REGION Network 2: Select with vacuum
   VAK:  NOP   0;
         SET;
         =     #OUT_H_Vacuum_active;
   //
         AN    #IN_P_Vacuum;
         L     S5T#500MS;
         SD    #IN_Timer_delay_Lock;
   //
         A     #IN_P_Vacuum;
         L     S5T#500MS;
         SD    #IN_Timer_delay_Pumpe;
   //
         AN    #IN_P_Vacuum;
         A     #IN_Timer_delay_Lock;
         =     #OUT_V_Lock_Vacuum;
   //
         ON    #IN_P_Vacuum;
         ON    #IN_Timer_delay_Pumpe;
         =     #OUT_V_Pump_Vacuum;
   //
         L     1;
         T     #IO_Status.Status_Vacuum;
END_REGION
END_FUNCTION

FUNCTION "FC107_Binär->Bit" : Void   // FC107, STL
TITLE = Chang a bin value in a bitcodetd value
{ S7_Optimized_Access := 'FALSE' }
AUTHOR : KT242
FAMILY : RS_KK
NAME : BintoBit
VERSION : 1.0
   VAR_INPUT
      IN_BinaerZahl : Byte;   // Eingabe einer Zahl (Maximal 16) als Ganzzahl
   END_VAR
   VAR_OUTPUT
      OUT_BitZahl : Word;   // Ausgabe der Zahl als Bitcodiertes Word
   END_VAR
   VAR_TEMP
      Temp_Sprungzaehler : Word;   // Zwischenmerker für einen Schleifenzähler
      Temp_Out_BitZahl : Word;
   END_VAR
BEGIN

REGION Network 1
         L     0;
         T     #Temp_Out_BitZahl;
   //
         O(;
         L     16;
         L     #IN_BinaerZahl;
         <I;
         );
         O(;
         L     1;
         <I;
         );
         JC    ENDE;
   //
         L     1;
         T     #Temp_Out_BitZahl;
   //
         L     #IN_BinaerZahl;
         ==I;
         JC    ENDE;
         L     1;
         -I;
   //
   NEXT: NOP   0;
         T     #Temp_Sprungzaehler;
   //
         L     #Temp_Out_BitZahl;
         SLW   1;
         T     #Temp_Out_BitZahl;
   //
         L     #Temp_Sprungzaehler;
         LOOP  NEXT;
   ENDE: NOP   0;

         L     #Temp_Out_BitZahl;
         T     #OUT_BitZahl;
END_REGION
END_FUNCTION

FUNCTION "FC111_FIFO" : Void   // FC111, STL
TITLE = FIFO of interface numbers
{ S7_Optimized_Access := 'FALSE' }
AUTHOR : KT242
FAMILY : RS_KK
NAME : FIFO
VERSION : 1.0
   VAR_INPUT
      IN_Amount_Interfaces : Int;   // Amount of interfaces to start shotcycle
      IN_Register : "UDT001_DWord_1_32";   // Data area of registered interfaces
      IN_Reset_List : Bool;   // Reset of list by new start of plc
      IN_StartAdr : Pointer;   // Start-addresse at DB to save countervalues to find out position at FIFO
      IN_DataBlock : DB_ANY;   // Datablock to save countervalues to find out position at FIFO
   END_VAR
   VAR_IN_OUT
      IO_FIRST : Int;   // Number of the member at first positon
      IO_SECOND : Int;   // Number of the member at second positon
      IO_FlagNewPos : Bool;   // Flag determine new positions at fifo
   END_VAR
   VAR_TEMP
      Schleifengroesse : Int;   // Schleifenzähler für den Durchlauf der Positionen bis "IN_Anzahl_Teilnehmer"
      Aktueller_Wert : Word;   // Wert des Zähler der eingetragenen Schnittstelle zur Erkennung der Position
      Wert_First : Word;   // Wert des Zähler der am längsten (first) eingetragenen Schnittstelle
      Wert_Second : Word;   // Wert des Zähler der am nächsten (second) eingetragenen Schnittstelle
      Baustein_Nr : Int;   // Merker zur Erkennung des Speicherbereiches der Bits "IN_Eintragen"
      Adresse_im_Baustein : DWord;   // and the start adress within the program block
      Eintragen_lokal : DWord;   // Zwischenspeicher der eingetragenen Formträgerschnittstellen (von UDT auf DWORD)
   END_VAR
BEGIN

REGION Network 1: FIFO - buffer
   // Am Ausgang "FIRST" liegt die Nummer des ersteingetragenen und an "SECOND" die 
   // des nachfolgenden Teilnehmers (max. 16) an. 
   // Am Eingangswort "Eintragen" muß das entsprechende Bit solange TRUE sein, bis
   // der Teilnehmer wieder ausgetragen werden kann.
   // Das Austragen des Teilnehmers erfolgt, wenn sich dieser in der Position "FIRST" 
   // oder "SECOND" befindet, innerhalb des Bausteins für die Schnittstelle.
   //_______________________________________________________________
   // Schieben der Eingetragenen FTs auf lokalen DWord- Bereich
   //
         L;
         LAR1;
         L     W[AR1, P#0.0];
         T     #Baustein_Nr;
   //
         L     D[AR1, P#2.0];
         T     #Adresse_im_Baustein;
         LAR2;
         L;
         LAR1;
   //
         OPN   DB[ #Baustein_Nr];
         L     DBD[AR2, P#0.0];
         T     LD[AR1, P#0.0];
   //__________________________________________________________
   //
         L     0;
         T     #Schleifengroesse;
         T     #Wert_First;
         T     #Wert_Second;
         L;
         LAR2;
   //
         L     #Eintragen_lokal;
         CAD;
         T     #Eintragen_lokal;
   //
         L;
         LAR1;
   //
         A(;
         L     #Eintragen_lokal;
         L     0;
         <>D;
         );
         JC    NEXT;
   //
   NEXT: A     "Flag_02_500_Hertz";
         FP    #IO_FlagNewPos;
         JCN   ENDE;
   //
         L     0;
         T     #IO_FIRST;
         T     #IO_SECOND;
   //
   M002: A     [AR1, P#0.0];  // Eintragebit ist gesetzt
         JCN   M001;
   //
         OPN   #IN_DataBlock;
         L     DBW[AR2, P#0.0];  // Speicherwert für eingetragene Station
         +     1;  // um 1 erhöhen
         T     DBW[AR2, P#0.0];
         T     #Aktueller_Wert;
   //
         L     #Aktueller_Wert;  // Wenn Speicherwert grösser als Maximum ist
         L     #Wert_First;
         >I;
         JCN   M011;
   //
         L     #Wert_First;
         T     #Wert_Second;
   //
         L     #Aktueller_Wert;  // Speicherwert in Maximum übertragen
         T     #Wert_First;
   //
         L     #IO_FIRST;
         T     #IO_SECOND;
   //
         L     #Schleifengroesse;  // Nummer der ersteingetragenen Station
         +     1;
         T     #IO_FIRST;
   //
         JU    M001;
   //
   M011: NOP   0;
         L     #Aktueller_Wert;  // Wenn Speicherwert grösser als Maximum ist
         L     #Wert_Second;
         >I;
         JCN   M001;
   //
         L     #Aktueller_Wert;  // Speicherwert in Maximum übertragen
         T     #Wert_Second;
   //
         L     #Schleifengroesse;  // Nummer der ersteingetragenen Station
         +     1;
         T     #IO_SECOND;
   //
   M001: A     [AR1, P#0.0];  // Eintragebit ist gesetzt
         JC    M003;
         L     0;  // wenn nicht gesetzt, dann ablöschen
         OPN   #IN_DataBlock;
         T     DBW[AR2, P#0.0];
   //
   M003: L     #Schleifengroesse;
         +     1;
         T     #Schleifengroesse;  // nächste Station
         +AR1  P#0.1;
         +AR2  P#2.0;
         L     #Schleifengroesse;  // Schleife ausführen,
         L     #IN_Amount_Interfaces;  // bis zur Anzahl der Teilnehmer
         <I;
         JC    M002;
   //
   ENDE: NOP   0;
END_REGION
END_FUNCTION

FUNCTION "FC112_IF_SP_MC" : Void   // FC112, STL
TITLE = Interface to switch panel and mould carrier
{ S7_Optimized_Access := 'FALSE' }
AUTHOR : KT242
FAMILY : RS_KK
NAME : SS_FT
VERSION : 1.4
// Function block to book in interface-no. of a foaming cycle by operation panel 
// or mould carrier interface.
   VAR_INPUT
      IN_InterfaceNo : Int;   // Number of related Interface
      IN_PositionFIRST : Int;   // No of interface, which is at first position // from FC 111 FIFO
      IN_PositionSECOND : Int;   // No of interface, which is at second position // from FC 111 FIFO
      IN_BCDSwitchPrgrNo_MH : Byte;   // Inputbyte of program no. from program selection switch at mixinghead panel
      IN_MH_Automatic : Bool;   // Mode switch mixing head panel at position cycle start "Auto"
      IN_MH_Manual : Bool;   // Mode switch mixing head panel at position cycle start "Manual"
      IN_Start_MH_Panel : Bool;   // Button start cycle at mixing head panel to enter interface no. -> FIFO
      IN_Stop_MH_Panel : Bool;   // Button stop cycle at mixing head panel to erase interface no. -> FIFO
      IN_ResetFault : Bool;   // Quit fault within this function block
      IN_ReleaseSWU : Bool;   // Switch over unit (SWU) of this interface is released
      IN_ReleaseMouldcarrier : Bool;   // Foaming release of mouldcarrier to enter interface number -> FIFO
      IN_PrgNoSwitchDeselected : Bool;   // Signal to bridge program selection by program selection switch
      IN_ReleaseFoaming : Bool;   // External signal release entering interface number
      IN_ReleaseCycle : Bool;   // Release start foaming cycle from function block cycle is active
      IN_OperationModeAuto : Bool;   // Foaming machine in automatic mode
      IN_OperationModeTest : Bool;   // Foaming machine in test mode; no foaming over mixinghead
      IN_LampTest : Bool;   // Check indicator lamp selected
      IN_CycleRunning : Bool;   // Foaming cycle is active
      IN_ShotRunning : Bool;   // Foaming active
      IN_LastStandbyTimeCycle : Bool;   // Last shot of foaming cycle was carried out
      IN_PulseCycleFinished : Bool;   // Pulse foaming cycle finished
   END_VAR
   VAR_OUTPUT
      OUT_Fault_To_MC : Bool;   // Output fault happend at active interface
      OUT_ShotEnd_To_MC : Bool;   // Output all part shots finished at this interface
      OUT_H_MH_Panel : Bool;   // Indicator foaming release and state of foaming cycle at mixinghead panel
   END_VAR
   VAR_IN_OUT
      IO_InterfaceActiveFIFO : Bool;   // Information interface no. active at FIFO
      IO_Status : "UDT112_IF_UP_MC";
      IO_Fault : "UDT1816_FLT_IF_SP_MC";
      IO_NewFault : Bool;
      IO_FaultLevel_1 : Bool;
      IO_FaultLevel_3 : Bool;
   END_VAR
   VAR_TEMP
      Temp_IO_Status : "UDT112_IF_UP_MC";
      TEMP_IO_Fault : "UDT1816_FLT_IF_SP_MC";
      Temp_ERROR_CODE : Int;   // Error state of systemfunction "BLKMOV" Blockmove
      AnyPointer1 : ANY;   // Pointer to copy thr array "IO_Status" and "Temp_IO_Status"
      AnyPointer2 : ANY;   // Pointer to copy thr array "IO_Status" and "Temp_IO_Status"
      Temp_SelectionPrgNo_OK : Bool;   // Flag selction program no. is OK at mixing head panel
      Temp_Flag_RelInterface : Bool;   // Flag release interface to enter at FIFO
      Temp_Pulse_RelInterface : Bool;   // Pulse für enter interface no. at FIFO
      Temp_Interface_at_Pos_1 : Bool;   // Flag interface at first position at FIFO
      Temp_Interface_at_Pos_2 : Bool;   // Flag interface at second position at FIFO
      Temp_Interface_Deselect : Bool;   // Flag deselct interface at FIFO
      Temp_Value_1 : Word;   // Value to calculate view between FUP/ KOP
      Temp_Value_2 : Int;   // Value to calculate view between FUP/ KOP
   END_VAR
BEGIN

REGION Network 1: Saved data integration
   // Änderungen:
   // -------------------------------------------------------------------------------
   // Anpassung der Aufschlüsselung der Schnittstellenstörungen.
   // v.d.Geest     20.09.2005
   // -------------------------------------------------------------------------------
   // Bei einer Störung der Gruppe 1 oder bei den zurücknehmen der Schäumfreigabe 
   // wird nur noch die Schnittstelle an der Position 1 ausgetragen.
   // (Änderungen auch im UDT112)
   // v.d.Geest     29.11.2004
   // -------------------------------------------------------------------------------
   // Genauere Aufschlüsselung der Schnittstellenstörungen. (Änderungen auch im 
   // UDT112)
   // Lindner       12.07.2004
   // -------------------------------------------------------------------------------
   // Bei Anwahl der Betriebsart "Testen" wird die Anzeigen der Schäumfreigabe an dem 
   // Bedienpult nicht mehr angezeigt.
   // Bereits vor dem einschalten der Betriebsart "Testen" eingetragene 
   // Schnittstellen werden noch bearbeitet, es können aber keine neuen eingetragen 
   // werden.
   // v.d.Geest     08.04.2003
   // -------------------------------------------------------------------------------
   // Das Signal "OUT_Schussende_an_FT" wurde über das Signal nach Ablauf der 
   // Kreislaufzeit 2 gebildet. Hierdurch konnte es vorkommen das sich mehrere 
   // Formträger die sich zum Schäumen angemeldet haben innerhalb eines Ablaufs der 
   // KLZ 2 abmelden. (Änderungen auch im UDT112)
   // v.d.Geest     17.03.2003
   // -------------------------------------------------------------------------------
   //-----
         LAR1;
         L;
         LAR2;
   //-----
         L     16#1002;  // Bytes
         T     W[AR1, P#0.0];
         L     2;  // Amount of bytes
         T     W[AR1, P#2.0];
         L     W[AR2, P#0.0];  // Block no,
         T     W[AR1, P#4.0];
         L     D[AR2, P#2.0];  // Startadress of datas
         T     D[AR1, P#6.0];
   //-----
         CALL  BLKMOV
         ( SRCBLK  := #AnyPointer1,
           RET_VAL := #Temp_ERROR_CODE,
           DSTBLK  := #Temp_IO_Status
         );
   //-----
         LAR1;
         L;
         LAR2;
   //-----
         L     16#1002;  // Bytes
         T     W[AR1, P#0.0];
         L     2;  // Amount of bytes
         T     W[AR1, P#2.0];
         L     W[AR2, P#0.0];  // Block no,
         T     W[AR1, P#4.0];
         L     D[AR2, P#2.0];  // Startadress of datas
         T     D[AR1, P#6.0];
   //-----
         CALL  BLKMOV
         ( SRCBLK  := #AnyPointer2,
           RET_VAL := #Temp_ERROR_CODE,
           DSTBLK  := #TEMP_IO_Fault
         );
   //-----
END_REGION

REGION Network 2: Test the program / program no. OK
   // Eine Schäumfreigabe über diese Schnittstelle darf nur erfolgen, wenn die 
   // Programmvorwahl ok ist. Dieses ist im Handbetrieb der Fall, sobald eine gültige 
   // Programmnummer an dem Wahlschalter des Mischkopfbedienpultes eingestellt wurde.
   //-----
         A(;
         A(;
         A(;
         L     #IN_BCDSwitchPrgrNo_MH;
         T     #Temp_Value_1;
         SET;
         SAVE;
         CLR;
         A     BR;
         );
         JNB   _001;
         L     #Temp_Value_1;
         L     16#FF;
         AW;
         T     #Temp_Value_1;
         SET;
         SAVE;
         CLR;
   _001: A     BR;
         );
         JNB   _002;
         L     #Temp_Value_1;
         T     #Temp_Value_2;
         SET;
         SAVE;
         CLR;
   _002: A     BR;
         );
         A(;
         L     #Temp_Value_2;
         L     0;
         <>I;
         );
         O     #IN_PrgNoSwitchDeselected;
         O(;
         A     #IN_CycleRunning;
         AN    #IN_Start_MH_Panel;
         AN    #IN_LastStandbyTimeCycle;
         );
         =     #Temp_SelectionPrgNo_OK;
END_REGION

REGION Network 3: Interface at position 1 of FIFO
         L     #IN_PositionFIRST;
         L     #IN_InterfaceNo;
         ==I;
         =     #Temp_IO_Status.IF_is_on_1_Position;
         =     #Temp_Interface_at_Pos_1;
END_REGION

REGION Network 4: Interface number to start next
         L     #IN_PositionSECOND;
         L     #IN_InterfaceNo;
         ==I;
         =     #Temp_IO_Status.IF_is_on_2_Position;
         =     #Temp_Interface_at_Pos_2;
END_REGION

REGION Network 5: Release mould carrier
         A(;
         A     #IN_MH_Automatic;
         A     #IN_ReleaseMouldcarrier;
         O     #IN_MH_Manual;
         );
         A     #Temp_SelectionPrgNo_OK;
         =     #Temp_Flag_RelInterface;
END_REGION

REGION Network 6: Sign out mouldcarrier by button Stop- foaming
         AN    #Temp_Interface_at_Pos_1;
         AN    #Temp_Interface_at_Pos_2;
         AN    #IN_Stop_MH_Panel;
         A     #IN_MH_Manual;
         S     #Temp_IO_Status.Stop_Buton_switched;
         A(;
         A     #IN_MH_Manual;
         A     #IN_Start_MH_Panel;
         A     #Temp_IO_Status.Stop_Buton_switched;
         ON    #Temp_IO_Status.IF_is_Selected;
         );
         R     #Temp_IO_Status.Stop_Buton_switched;
         NOP   0;
END_REGION

REGION Network 7: Fault at the interface
         A(;
         A(;
         ON    #IN_MH_Automatic;
         O     #IN_ResetFault;
         );
         R     #TEMP_IO_Fault.Fault_IF;

         A(;
         AN    #IN_MH_Manual;
         AN    #IN_MH_Automatic;
         O(;
         AN    #Temp_Flag_RelInterface;
         A     #IN_CycleRunning;
         AN    #IN_LastStandbyTimeCycle;
         );
         O(;
         A(;
         O     #IO_FaultLevel_1;
         ON    #IN_ReleaseFoaming;
         ON    #IN_ReleaseCycle;
         );
         FP    #Temp_IO_Status.FHF_Fault;
         AN    #IN_LastStandbyTimeCycle;
         A     #Temp_Interface_at_Pos_1;
         );
         ON    #IN_OperationModeAuto;
         ON    #IN_ReleaseSWU;
         O;
         A(;
         O     #Temp_Interface_at_Pos_1;
         O     #Temp_Interface_at_Pos_2;
         );
         A(;
         O     #Temp_IO_Status.Stop_Buton_switched;
         ON    #IN_Stop_MH_Panel;
         );
         );
         A     #Temp_IO_Status.IF_is_Selected;
         AN    #TEMP_IO_Fault.Fault_IF;
         S     #IO_NewFault;
         S     #TEMP_IO_Fault.Fault_IF;
         A     #TEMP_IO_Fault.Fault_IF;
         );
         A     #IN_MH_Automatic;
         =     #OUT_Fault_To_MC;
END_REGION

REGION Network 8: Shotend
         A(;
         A(;
         ON    #IN_MH_Automatic;
         O;
         AN    #Temp_Flag_RelInterface;
         AN    #TEMP_IO_Fault.Fault_IF;
         );
         R     #Temp_IO_Status.Shotsend_IF;
         A(;
         O     #TEMP_IO_Fault.Fault_IF;
         O     #IN_PulseCycleFinished;
         );
         FP    #Temp_IO_Status.FHF_KLZ2;
         A     #Temp_Interface_at_Pos_1;
         S     #Temp_IO_Status.Shotsend_IF;
         A     #Temp_IO_Status.Shotsend_IF;
         );
         A     #IN_MH_Automatic;
         =     #OUT_ShotEnd_To_MC;
END_REGION

REGION Network 9: Log in interface no at FIFO
         A(;
         A     #IN_Start_MH_Panel;
         FP    #Temp_IO_Status.HF_T_Start_MH;
         A     #IN_MH_Manual;
         O;
         A(;
         A     #IN_ReleaseMouldcarrier;
         BLD   100;
         FP    #Temp_IO_Status.HF_Release_IF;
         );
         A     #IN_MH_Automatic;
         );
         AN    #IN_OperationModeTest;
         A     #Temp_Flag_RelInterface;
         A     #IN_ReleaseSWU;
         A     #IN_ReleaseFoaming;
         A     #IN_ReleaseCycle;
         AN    #Temp_IO_Status.IF_is_Selected;
         AN    #Temp_IO_Status.Shotsend_IF;
         AN    #TEMP_IO_Fault.Fault_IF;
         S     #Temp_IO_Status.IF_is_Selected;
         S     #IO_InterfaceActiveFIFO;
END_REGION

REGION Network 10: Log off interface no. at FIFO
         A     #IN_PulseCycleFinished;
         A     #Temp_Interface_at_Pos_1;
         O;
         AN    #Temp_Flag_RelInterface;
         AN    #Temp_Interface_at_Pos_1;
         ON    #IN_OperationModeAuto;
         O     #TEMP_IO_Fault.Fault_IF;
         A     #Temp_IO_Status.IF_is_Selected;
         =     #Temp_Interface_Deselect;
         R     #Temp_IO_Status.IF_is_Selected;
         R     #IO_InterfaceActiveFIFO;
END_REGION

REGION Network 11: Start cycle with this interface
         A     #Temp_IO_Status.IF_is_Selected;
         A     #Temp_Interface_at_Pos_1;
         A     #IN_ReleaseFoaming;
         A     #IN_ReleaseCycle;
         AN    #IN_CycleRunning;
         =     #Temp_IO_Status.Start_to_Cycle;
END_REGION

REGION Network 12: Break cycle at this interface
         AN    #Temp_IO_Status.IF_is_Selected;
         A     #Temp_Interface_at_Pos_1;
         AN    #IN_LastStandbyTimeCycle;
         A     #IN_CycleRunning;
         =     #Temp_IO_Status.Stop_to_Cycle;
END_REGION

REGION Network 13: Set indicater ready for foaming
         A(;
         A     #Temp_Flag_RelInterface;
         A     #IN_MH_Manual;
         O     #IN_MH_Automatic;
         );
         A     #IN_ReleaseFoaming;
         A     #IN_ReleaseCycle;
         A(;
         ON    #Temp_IO_Status.Shotsend_IF;
         O;
         A     #IN_LastStandbyTimeCycle;
         A     #Temp_Interface_at_Pos_1;
         );
         A(;
         AN    #Temp_IO_Status.IF_is_Selected;
         A     #IN_MH_Manual;
         AN    #IN_OperationModeTest;
         O;
         A     #Temp_IO_Status.IF_is_Selected;
         A(;
         AN    #Temp_Interface_at_Pos_1;
         A     "Flag_00_500_Hertz";
         O;
         A     #Temp_Interface_at_Pos_1;
         A(;
         AN    #IN_ShotRunning;
         A     "Flag_01_000_Hertz";
         O;
         A     #IN_ShotRunning;
         A     "Flag_05_000_Hertz";
         );
         );
         );
         A     #Temp_SelectionPrgNo_OK;
         A     #IN_ReleaseSWU;
         AN    #TEMP_IO_Fault.Fault_IF;
         O     #IN_LampTest;
         =     #OUT_H_MH_Panel;
END_REGION

REGION Network 14: Reset of faults
         O     #IN_ResetFault;
         R     #TEMP_IO_Fault.FLT_pouring_release;
         R     #TEMP_IO_Fault.FLT_SWU_release;
         R     #TEMP_IO_Fault.FLT_Stop_while_selected;
         R     #TEMP_IO_Fault.FLT_op_mode_O;
         R     #TEMP_IO_Fault.FLT_Cycle_release;
END_REGION

REGION Network 15: Fault foaming release (external signal)
   // Störung: Die Schäumfreigebe wurde auf 0 gesetzt. Während der Formträger 
   // angemeldet und an erster Position ist.
   // - #Temp_IO_Status.Stoerung_Schaeumfreigabe -
         AN    #IN_ReleaseFoaming;
         AN    #IN_LastStandbyTimeCycle;
         A     #Temp_Interface_Deselect;
         A     #Temp_Interface_at_Pos_1;
         A     #IN_MH_Automatic;
         AN    #TEMP_IO_Fault.FLT_pouring_release;
         S     #IO_NewFault;
         S     #TEMP_IO_Fault.FLT_pouring_release;
END_REGION

REGION Network 16: Fault SWU release set to 0 (external signal)
   // Störung: Die USE-Freigabe wurde auf 0 gesetzt. Während der Formträger 
   // angemeldet ist.
   // - #Temp_IO_Status.USE_Freigabe-
         AN    #IN_ReleaseSWU;
         A     #Temp_Interface_Deselect;
         AN    #TEMP_IO_Fault.FLT_pouring_release;
         AN    #TEMP_IO_Fault.FLT_SWU_release;
         S     #IO_NewFault;
         S     #TEMP_IO_Fault.FLT_SWU_release;
END_REGION

REGION Network 17: Fault STOP-button pressed during foaming cycle
   // Störung: Der STOP-Taster wurde auf 0 gesetzt. Während der Formträger 
   // angemeldet und an erster Position ist.
   // -#Temp_IO_Status.Stoerung_STOP_Taster-
         A(;
         O     #Temp_Interface_at_Pos_1;
         O     #Temp_Interface_at_Pos_2;
         );
         A(;
         O     #Temp_IO_Status.Stop_Buton_switched;
         ON    #IN_Stop_MH_Panel;
         );
         A     #Temp_Interface_Deselect;
         AN    #TEMP_IO_Fault.FLT_pouring_release;
         AN    #TEMP_IO_Fault.FLT_SWU_release;
         AN    #TEMP_IO_Fault.FLT_Stop_while_selected;
         S     #IO_NewFault;
         S     #TEMP_IO_Fault.FLT_Stop_while_selected;
END_REGION

REGION Network 18: Fault key-switch manual/auto at MH-panel set to 0
   // Störung: Der Hand/Auto Schlüsselschalter wurde auf 0 gesetzt. Während der 
   // Formträger angemeldet und an erster Position ist.
   // -#Temp_IO_Status.Stoerung_Hand_Auto-
         AN    #IN_MH_Manual;
         AN    #IN_MH_Automatic;
         A     #Temp_Interface_at_Pos_1;
         AN    #TEMP_IO_Fault.FLT_pouring_release;
         AN    #TEMP_IO_Fault.FLT_SWU_release;
         AN    #TEMP_IO_Fault.FLT_Stop_while_selected;
         AN    #TEMP_IO_Fault.FLT_op_mode_O;
         S     #IO_NewFault;
         S     #TEMP_IO_Fault.FLT_op_mode_O;
END_REGION

REGION Network 19: Fault foaming release
   // Störung: Freigabe Zyklus wurde auf 0 gesetzt. Während der 
   // Formträger angemeldet und an erster Position ist.
         AN    #IN_ReleaseCycle;
         AN    #IN_LastStandbyTimeCycle;
         A     #Temp_Interface_at_Pos_1;
         AN    #TEMP_IO_Fault.FLT_pouring_release;
         AN    #TEMP_IO_Fault.FLT_SWU_release;
         AN    #TEMP_IO_Fault.FLT_Stop_while_selected;
         AN    #TEMP_IO_Fault.FLT_op_mode_O;
         AN    #TEMP_IO_Fault.FLT_Cycle_release;
         S     #IO_NewFault;
         S     #TEMP_IO_Fault.FLT_Cycle_release;
END_REGION

REGION Network 20: Error handling
         O     #TEMP_IO_Fault.FLT_pouring_release;
         O     #TEMP_IO_Fault.FLT_SWU_release;
         O     #TEMP_IO_Fault.FLT_Stop_while_selected;
         O     #TEMP_IO_Fault.FLT_op_mode_O;
         O     #TEMP_IO_Fault.FLT_Cycle_release;
         O     #TEMP_IO_Fault.Fault_IF;
         S     #IO_FaultLevel_3;
END_REGION

REGION Network 21: Save data
   //-----
         CALL  BLKMOV
         ( SRCBLK  := #Temp_IO_Status,
           RET_VAL := #Temp_ERROR_CODE,
           DSTBLK  := #AnyPointer1
         );
   //-----
         CALL  BLKMOV
         ( SRCBLK  := #TEMP_IO_Fault,
           RET_VAL := #Temp_ERROR_CODE,
           DSTBLK  := #AnyPointer2
         );
   //-----
END_REGION
END_FUNCTION

FUNCTION "FC114_IF_externalPlant" : Void   // FC114, STL
TITLE = Interface between machine and external plant
{ S7_Optimized_Access := 'FALSE' }
AUTHOR : KT242
NAME : SS_AP
VERSION : 1.1
   VAR_INPUT
      IN_Release : Bool;   // General release of interface external plant
      IN_use_Inv_Program : Bool;   // Number transfer by using an inverse program number
      IN_use_Parity_Bit : Bool;   // Number transfer by using parity check
      IN_Reset_fault_Fkt : Bool;   // Signal to reset faults at innerhalb this function block
      IN_Stop_MH_OpPanel : Bool;   // Stop- signal at MH - operator panel to put out interfacenumber from FIFO
      IN_Operationmode_Operate : Bool;   // Foaming machine in operation mode with foam dispersion
      IN_MH_panel_automatic : Bool;   // Mixinghead - operator panel switched to automatic
      IN_FCycleRelease_extern : Bool;   // Foaming release from externen plant
      IN_FCycle_release : Bool;   // Release start foaming cycle from function block cycle
      IN_FCycle_running : Bool;   // Foaming cycle is running
      IN_FCycle_Shotrelease : Bool;   // Foaming release from Schäumzyklus steht an
      IN_FCycle_Shot_running : Bool;   // Foaming happens
      IN_FCycle_Pulse_Shotend : Bool;   // Foaming finished
      IN_FCycle_Pulse_End : Bool;   // Pulse foaming cycle finished // Signal takes 1 SPS- Cycle
      IN_ExtPlant_OK : Bool;   // Signal from external plant: External plant is ready for production
      IN_Strobe_or_Start : Bool;   // Signal from external plant: Strobe valid or cycle start signal
      IN_StrobeINV_or_Parity : Bool;   // Signal from external plant: Data strobe inverse or parity bit
      IN_Start_Shot : Bool;   // Signal from external plant: Start foaming by shot release from PU
      IN_CP_forward : Bool;   // Signal from external plant: Trigger cleaning piston
      IN_ProgNo_ExtPlant : Byte;   // Signal from external plant: Program no or inverse program number
      IN_maxAmount_ProgNo : Int;   // Limitation of program number from external plant
   END_VAR
   VAR_OUTPUT
      OUT_PU_OK : Bool;   // Signal to external Plant: Foaming machine is ready to start foaming cycle
      OUT_Strobe_quit : Bool;   // Signal to external Plant: Program number (..Invers) was accepted
      OUT_FCycle_running : Bool;   // Signal to external Plant: Foaming cycle was started and runs
      OUT_ReadyForFoaming : Bool;   // Signal to external Plant: Foaming machine ready to open mixinghead
      OUT_FoamingActive : Bool;   // Signal to external Plant: Foaming is going on
      OUT_FoamingEnd : Bool;   // Signal to external Plant: Foaming is finished
      OUT_ServiceShot : Bool;   // Signal to external Plant: Foaming machine is at service mode
   END_VAR
   VAR_IN_OUT
      IO_Status : "UDT114_IF_externalPlant";
      IO_Fault : "UDT1817_FLT_IF_extPlant";
      IO_NewFault : Bool;
      IO_FaultLevel_1 : Bool;
      IO_FaultLevel_2 : Bool;
      IO_FaultLevel_3 : Bool;
   END_VAR
   VAR_TEMP
      Temp_IO_Status : "UDT114_IF_externalPlant";
      TEMP_IO_Fault : "UDT1817_FLT_IF_extPlant";
      ERROR_CODE : Int;   // Error state of systemfunction "BLKMOV" Blockmove
      AnyPointer1 : ANY;   // Pointer to copy thr array "IO_Status" and "Temp_IO_Status"
      AnyPointer2 : ANY;   // Pointer to copy thr array "IO_Status" and "Temp_IO_Status"
      Temp_ProgNo_Puls : Byte;   // Temporärer Zwischenspeicher der Programmnummer für die Paritätsprüfung
      Strobe_quitt_reset : Bool;   // Hilfsmerker zum zurücksetzen des Quittierungsbits
      Temp_PulseCycleRelease : Bool;   // Impulshilfsmerker das das starten einen Schäumzyklusses Freigegeben ist
      Temp_Pulse_ExtP_Start : Bool;   // Impulshilfsmerker für das Starten die Programmermittlung des Schnittstelle
   END_VAR
BEGIN

REGION Network 1: Saved data integration
   // Änderungen:
   // -------------------------------------------------------------------------------
   // Wenn beim starten der Anlage das Stobe Bit von der Fremdanlage schon oder noch 
   // gesetzt war wurde direkt ein Schäumprogramm gestartet.
   // Durch eine Flankenabfrage des Signals "#IN_Strobe_oder_Start" im Netzwerk 3 
   // wurde dieses unterbunden
   // 
   // Jäger       19.08.2004
   // -------------------------------------------------------------------------------
   //-----
         LAR1;
         L;
         LAR2;
   //-----
         L     16#1002;  // Bytes
         T     W[AR1, P#0.0];
         L     6;  // Amount of bytes
         T     W[AR1, P#2.0];
         L     W[AR2, P#0.0];  // Block no,
         T     W[AR1, P#4.0];
         L     D[AR2, P#2.0];  // Startadress of datas
         T     D[AR1, P#6.0];
   //-----
         CALL  BLKMOV
         ( SRCBLK  := #AnyPointer1,
           RET_VAL := #ERROR_CODE,
           DSTBLK  := #Temp_IO_Status
         );
   //-----
         LAR1;
         L;
         LAR2;
   //-----
         L     16#1002;  // Bytes
         T     W[AR1, P#0.0];
         L     2;  // Amount of bytes
         T     W[AR1, P#2.0];
         L     W[AR2, P#0.0];  // Block no,
         T     W[AR1, P#4.0];
         L     D[AR2, P#2.0];  // Startadress of datas
         T     D[AR1, P#6.0];
   //-----
         CALL  BLKMOV
         ( SRCBLK  := #AnyPointer2,
           RET_VAL := #ERROR_CODE,
           DSTBLK  := #TEMP_IO_Fault
         );
   //-----
END_REGION

REGION Network 2: Reset and set of faults
         CLR;
         =     #Temp_IO_Status.FaultLevel_1;
         =     #Temp_IO_Status.FaultLevel_2;
         =     #Temp_IO_Status.FaultLevel_3;
         =     #Temp_IO_Status.Message_activ;
   //-----
         A     #IN_Reset_fault_Fkt;
         R     #TEMP_IO_Fault.FLT_Strobe;
         R     #TEMP_IO_Fault.FLT_Strobe_inv;
         R     #TEMP_IO_Fault.FLT_AP_not_OK;
         R     #TEMP_IO_Fault.FLT_no_number;
         R     #TEMP_IO_Fault.FLT_inverse_number;
         R     #TEMP_IO_Fault.FLT_Parity_Bit;
         R     #TEMP_IO_Fault.FLT_Cycle_Stoped;
         R     #TEMP_IO_Fault.FLT_Start_Shot;
   //
         O     #IN_FCycle_release;
         FP    #Temp_IO_Status.FHF_Cycle_Release;
         =     #Temp_PulseCycleRelease;
   //
         O     #Temp_PulseCycleRelease;
         ON    #IN_ExtPlant_OK;
         A     #IN_Strobe_or_Start;
         A     #IN_MH_panel_automatic;
         AN    #TEMP_IO_Fault.FLT_Start_Shot;
         AN    #TEMP_IO_Fault.FLT_no_number;
         AN    #TEMP_IO_Fault.FLT_Strobe;
         S     #TEMP_IO_Fault.FLT_Strobe;
         S     #IO_NewFault;
   //
         O     #Temp_PulseCycleRelease;
         ON    #IN_ExtPlant_OK;
         A     #IN_StrobeINV_or_Parity;
         AN    #IN_use_Parity_Bit;
         A     #IN_MH_panel_automatic;
         AN    #TEMP_IO_Fault.FLT_no_number;
         AN    #TEMP_IO_Fault.FLT_Strobe_inv;
         S     #TEMP_IO_Fault.FLT_Strobe_inv;
         S     #IO_NewFault;
   //
         A     #IN_ExtPlant_OK;
         A     #IN_FCycle_release;
         A     #IN_Start_Shot;
         A     #IN_Strobe_or_Start;
         A     #IN_MH_panel_automatic;
         AN    #Temp_IO_Status.PU_Shotend;
         AN    #Temp_IO_Status.IF_is_selected;
         AN    #TEMP_IO_Fault.FLT_Start_Shot;
         S     #TEMP_IO_Fault.FLT_Start_Shot;
         S     #IO_NewFault;
   //
         AN    #IN_ExtPlant_OK;
         A     #IN_Release;
         A     #IN_MH_panel_automatic;
         AN    #TEMP_IO_Fault.FLT_AP_not_OK;
         =     #TEMP_IO_Fault.MSG_AP_not_OK;
         S     #Temp_IO_Status.Message_activ;
   //
         AN    #IN_ExtPlant_OK;
         A     #IN_Release;
         A     #IN_FCycle_release;
         A     #IN_MH_panel_automatic;
         AN    #TEMP_IO_Fault.FLT_AP_not_OK;
         S     #TEMP_IO_Fault.FLT_AP_not_OK;
         S     #IO_NewFault;
   //
END_REGION

REGION Network 3: Raising edge of Start/ Strobe- signal
         A     #IN_Strobe_or_Start;
         FP    #Temp_IO_Status.HF_StrobeStart;
         =     #Temp_Pulse_ExtP_Start;
END_REGION

REGION Network 4: Release start signal detection
         A     #IN_FCycle_release;
         A     #IN_Release;
         A     #IN_ExtPlant_OK;
         A     #IN_Stop_MH_OpPanel;
         A     #IN_MH_panel_automatic;
         AN    #TEMP_IO_Fault.FLT_Strobe;
         AN    #TEMP_IO_Fault.FLT_Strobe_inv;
         AN    #TEMP_IO_Fault.FLT_Start_Shot;
         AN    #TEMP_IO_Fault.FLT_AP_not_OK;
         AN    #TEMP_IO_Fault.FLT_Parity_Bit;
         AN    #TEMP_IO_Fault.FLT_Cycle_Stoped;
         JCN   res;
END_REGION

REGION Network 5: Select signal transver mode (Invers or Parity)
   // Dieser Baustein kann wahlweise für verschiedene Fremdanlagenschnittstellen 
   // verwendet werden.
   // - Hardwareschnittstelle mit Programm und invertiertem Programm
   // - Profibusschnittstelle nur mit einer Programmnummer
   // - Schnittstelle mit Paritätsbitüberbrüfung
         A     #IN_use_Parity_Bit;
         JC    PaCh;  // Jump to parity check
END_REGION

REGION Network 6: Sprungleiste fuer Invers check
         L     #Temp_IO_Status."Step";
         JL    res1;
         JU    stro;  // case 0     Strobe
         JU    qstr;  // case 1     quitt Strobe
         JU    istr;  // case 2     Strobe invers
         JU    qist;  // case 3     quitt Strobe invers
         JU    wait;  // case 4     Wait till Null
   //
   res1: JU    res;
END_REGION

REGION Network 7: Strobe
   stro: NOP   0;
         A     #Temp_Pulse_ExtP_Start;  //Edge Strobe or Start signal
         JCN   ausg;
   //
         A(;
         L     #IN_ProgNo_ExtPlant;
         L     0;
         <=I;
         );
         A(;
         L     #IN_ProgNo_ExtPlant;
         L     #IN_maxAmount_ProgNo;
         >I;
         );
         AN    #TEMP_IO_Fault.FLT_no_number;
         S     #TEMP_IO_Fault.FLT_no_number;
         S     #IO_NewFault;
   //
         L     #IN_ProgNo_ExtPlant;
         T     #Temp_IO_Status.PrgNo_Storage;
   //
         A     #IN_use_Inv_Program;
         JC    J_qu;
   //
         L     3;
         T     #Temp_IO_Status."Step";
         JU    ausg;
   //
   J_qu: L     1;
         T     #Temp_IO_Status."Step";
   //
         JU    ausg;
END_REGION

REGION Network 8: Confirme strobe
   qstr: NOP   0;  // case 1
         A     #IN_Strobe_or_Start;
         S     #OUT_Strobe_quit;
   //
         AN    #IN_Strobe_or_Start;
         A     #OUT_Strobe_quit;
         R     #OUT_Strobe_quit;
         JCN   ausg;
         L     2;
         T     #Temp_IO_Status."Step";
         JU    ausg;
END_REGION

REGION Network 9: Strobe invers und check ob ok
   istr: NOP   0;  // case 2
         A     #IN_StrobeINV_or_Parity;
         JCN   ausg;
         L     #IN_ProgNo_ExtPlant;
         L     #Temp_IO_Status.PrgNo_Storage;
         +I;
         L     255;
         ==I;
         NOT;
         AN    #TEMP_IO_Fault.FLT_inverse_number;
         S     #TEMP_IO_Fault.FLT_inverse_number;
         S     #IO_NewFault;
   //
         L     3;
         T     #Temp_IO_Status."Step";
   //
         JU    ausg;
END_REGION

REGION Network 10: Confirm (Quitt) strobe invers
   qist: NOP   0;  // case 3
   //
         A     #IN_StrobeINV_or_Parity;
         A     #IN_use_Inv_Program;
         O     #IN_Strobe_or_Start;
         S     #OUT_Strobe_quit;
   //
         L     4;
         T     #Temp_IO_Status."Step";
   //
         AN    #TEMP_IO_Fault.FLT_no_number;
         AN    #TEMP_IO_Fault.FLT_inverse_number;
         S     #Temp_IO_Status.IF_is_selected;
   //
         JU    ausg;
END_REGION

REGION Network 11: Warte auf strobe/ strobe invers auf Null
   wait: NOP   0;  // case 4
   //
         A     #IN_StrobeINV_or_Parity;
         A     #IN_use_Inv_Program;
         O     #IN_Strobe_or_Start;
         JC    Next;
         L     0;
         T     #Temp_IO_Status."Step";
         SET;
         R     #OUT_Strobe_quit;
   //
   Next: NOP   0;
   //
         JU    ausg;  // Jump over Parity check
END_REGION

REGION Network 12: Parity Check
   PaCh: NOP   0;
   //
         A     #Temp_Pulse_ExtP_Start;
         AN    #Temp_IO_Status.IF_is_selected;
         JCN   ausg;
   //
         L     #IN_ProgNo_ExtPlant;
         T     #Temp_ProgNo_Puls;
         T     #Temp_IO_Status.PrgNo_Storage;
   //
         X     #Temp_ProgNo_Puls.%X0;
         X     #Temp_ProgNo_Puls.%X1;
         X     #Temp_ProgNo_Puls.%X2;
         X     #Temp_ProgNo_Puls.%X3;
         X     #Temp_ProgNo_Puls.%X4;
         X     #Temp_ProgNo_Puls.%X5;
         X     #Temp_ProgNo_Puls.%X6;
         X     #Temp_ProgNo_Puls.%X7;
         X     #IN_StrobeINV_or_Parity;
         S     #TEMP_IO_Fault.FLT_Parity_Bit;
         S     #IO_NewFault;

   //
         O(;
         L     0;
         L     #Temp_ProgNo_Puls;
         >=I;
         );
         O(;
         L     #IN_maxAmount_ProgNo;
         >I;
         );
         S     #TEMP_IO_Fault.FLT_no_number;
         S     #IO_NewFault;
   //
         AN    #TEMP_IO_Fault.FLT_Parity_Bit;
         AN    #TEMP_IO_Fault.FLT_no_number;
         S     #Temp_IO_Status.IF_is_selected;
   //
         JU    ausg;
END_REGION

REGION Network 13: Reset
   res:  NOP   0;
         A     #Temp_IO_Status.IF_is_selected;
         =     #Temp_IO_Status.Stop_to_Cycle;
   //     UN    #TEMP_IO_Fault.FLT_Cycle_Stoped
   //      S     #TEMP_IO_Fault.FLT_Cycle_Stoped
   //      S     #IO_NewFault
   //
         SET;
         R     #Temp_IO_Status.IF_is_selected;
         R     #OUT_Strobe_quit;
         R     #Temp_IO_Status.Start_to_Cycle;
         R     #Temp_IO_Status.ExtP_MH_open;
         R     #Temp_IO_Status.ExtP_CP_forward;
   //
         A     #IN_StrobeINV_or_Parity;
         O     #IN_Strobe_or_Start;
         =     #OUT_Strobe_quit;
   //
         L     0;
         T     #Temp_IO_Status."Step";
         T     #Temp_IO_Status.PrgNo_Storage;
END_REGION

REGION Network 14: Starten des Schäumzyklusses
   ausg: NOP   0;
   //
         A     #Temp_IO_Status.IF_is_selected;
         AN    #IN_FCycle_running;
         =     #Temp_IO_Status.Start_to_Cycle;
         JCN   shot;
   //
         L     #Temp_IO_Status.PrgNo_Storage;
         T     #Temp_IO_Status.PrgNo_to_PU;
   //
   shot: NOP   0;
   //
         O     #IN_FCycle_Pulse_End;
         JCN   Goon;
   //
         SET;
         R     #Temp_IO_Status.IF_is_selected;
         L     0;
         T     #Temp_IO_Status.PrgNo_to_PU;
   //
   Goon: NOP   0;
END_REGION

REGION Network 15: Bilden der Signale an die/ von der Fremdanlage
   //______________________________________________
   // Die Schäummaschine ist Betriebsbereit
   //
         A     #IN_Release;
         A     #IN_FCycle_release;
         A     #IN_MH_panel_automatic;
         =     #Temp_IO_Status.PU_ok;
   //
         A     #IN_FCycle_running;
         A     #IN_MH_panel_automatic;
         =     #Temp_IO_Status.PU_Cycle_runs;
   //______________________________________________
   // Freigabe zum Ansteuern des Mischkofes
   //
         A     #IN_FCycle_Shotrelease;
         AN    #Temp_IO_Status.PU_Shotend;
         =     #Temp_IO_Status.PU_Pouringrelease;
   //______________________________________________
   // Bilden des Signal Schuss beendet
   //
         A     #IN_FCycle_Pulse_Shotend;
         S     #Temp_IO_Status.PU_Shotend;
   //
         AN    #IN_Start_Shot;
         A     #Temp_IO_Status.PU_Shotend;
         S     #Temp_IO_Status.StatShotOffafterCycleFinish;
         AN    #IN_FCycle_running;
         A     #Temp_IO_Status.PU_Shotend;
         S     #Temp_IO_Status.CycleOffafterShotFinish;
   //
         A     #Temp_IO_Status.StatShotOffafterCycleFinish;
         A     #Temp_IO_Status.CycleOffafterShotFinish;
         R     #Temp_IO_Status.PU_Shotend;
         R     #Temp_IO_Status.StatShotOffafterCycleFinish;
         R     #Temp_IO_Status.CycleOffafterShotFinish;
   //______________________________________________
   // Ansteuern des Mischkopfventils von der Fremdanlage
   //
         A     #IN_Start_Shot;
         A     #IN_FCycle_running;
         A     #IN_MH_panel_automatic;
         AN    #Temp_IO_Status.PU_Shotend;
         =     #Temp_IO_Status.ExtP_MH_open;
   //______________________________________________
   // Ansteuern des Reinigungskolben von der Fremdanlage
   //
         A     #IN_CP_forward;
         =     #Temp_IO_Status.ExtP_CP_forward;
   //______________________________________________
   // Signal das sich die Fremdanlage im Automatikbetrieb befindet
   //
         A     #IN_ExtPlant_OK;
         =     #Temp_IO_Status.ExtP_in_Automatic;
END_REGION

REGION Network 16: Ansteuern der Signale an die Fremdanlage
         A     #Temp_IO_Status.PU_ok;
         =     #OUT_PU_OK;
   //
         A     #Temp_IO_Status.PU_Cycle_runs;
         =     #OUT_FCycle_running;
   //
         A     #IN_FCycle_Shot_running;
         =     #OUT_FoamingActive;
   //
         A     #Temp_IO_Status.PU_Pouringrelease;
         =     #OUT_ReadyForFoaming;
   //
         A     #Temp_IO_Status.PU_Shotend;
         =     #OUT_FoamingEnd;
   //
         AN    #IN_Operationmode_Operate;
         =     #OUT_ServiceShot;
END_REGION

REGION Network 17: Error handling
   //      O     XXXXXXXX
   //      S     #Temp_IO_Status.FaultLevel_1
   //      S     #IO_FaultLevel_1

   //      O     XXXXXXXX
   //      S     #Temp_IO_Status.FaultLevel_2
   //      S     #IO_FaultLevel_2

         O     #TEMP_IO_Fault.FLT_Strobe;
         O     #TEMP_IO_Fault.FLT_Strobe_inv;
         O     #TEMP_IO_Fault.FLT_AP_not_OK;
         O     #TEMP_IO_Fault.FLT_no_number;
         O     #TEMP_IO_Fault.FLT_inverse_number;
         O     #TEMP_IO_Fault.FLT_Parity_Bit;
         O     #TEMP_IO_Fault.FLT_Cycle_Stoped;
         O     #TEMP_IO_Fault.FLT_Start_Shot;
         S     #Temp_IO_Status.FaultLevel_3;
         S     #IO_FaultLevel_3;
END_REGION

REGION Network 18: Save data
         CALL  BLKMOV
         ( SRCBLK  := #Temp_IO_Status,
           RET_VAL := #ERROR_CODE,
           DSTBLK  := #AnyPointer1
         );
   //
         CALL  BLKMOV
         ( SRCBLK  := #TEMP_IO_Fault,
           RET_VAL := #ERROR_CODE,
           DSTBLK  := #AnyPointer2
         );
   //
END_REGION
END_FUNCTION

FUNCTION "FC115_Testen" : Void   // FC115, STL
TITLE = Halbautomatisches Testen über Ventile
{ S7_Optimized_Access := 'FALSE' }
AUTHOR : KT242
FAMILY : RS_KK
NAME : Testen
VERSION : 1.1
   VAR_INPUT
      IN_Betriebsart_Testen : Bool;   // Die Schäummaschine befindet sich in der Betriebsart Testen über Ventil
      IN_Betriebsart_Betrieb : Bool;   // Die Schäummaschine befindet sich im der Betriebsart mit Schaumaustrag
      IN_Lampentest : Bool;   // Zur Überprüfung der Anzeigen wurde ein Lampentest angewählt
      IN_Start_Testen_K1 : Bool;   // Taster zum Starten der Testfunktion für Komponente 01
      IN_Start_Testen_K2 : Bool;   // Taster zum Starten der Testfunktion für Komponente 02
      IN_Start_Testen_K3 : Bool;   // Taster zum Starten der Testfunktion für Komponente 03
      IN_Start_Testen_K4 : Bool;   // Taster zum Starten der Testfunktion für Komponente 04
      IN_Stop_Testen : Bool;   // Taster zum Stoppen aller aktuellen Testfunktionen
      IN_Stoerung_Gruppe_1 : Bool;   // Eine Störung der Gruppe 1 steht an und wurde noch nicht quittiert
      IN_Zyklus_Freigabe : Bool;   // Die Freigabe zum Starten des Schäumzyklusses aus dem Zyklusbaustein steht an
      IN_Zyklus_laeuft : Bool;   // Ein Schäumzyklus wurde bereits gestartet
      IN_Zyklus_Schuss_laeuft : Bool;   // Der im Schäumprogramm eingegebene Austrag wird durchgeführt
      IN_Imp_Zyklus_Ende : Bool;   // Der Schäumzyklus wurde beendet // Signal für 1 SPS- Zyklus
      IN_Zyklus_KLZ2_u_ff : Bool;   // Der letzte Teilschuß des Schäumprogramms wurde ausgeführt
   END_VAR
   VAR_OUTPUT
      OUT_H_Testen_K1 : Bool;   // Anzeige des Zustandes der Testfunktion der Komponente 1
      OUT_H_Testen_K2 : Bool;   // Anzeige des Zustandes der Testfunktion der Komponente 2
      OUT_H_Testen_K3 : Bool;   // Anzeige des Zustandes der Testfunktion der Komponente 3
      OUT_H_Testen_K4 : Bool;   // Anzeige des Zustandes der Testfunktion der Komponente 4
      OUT_V_Testen_K1 : Bool;   // Ansteuerung des Rücklaufventils zum Testen der Komponente 1
      OUT_V_Testen_K2 : Bool;   // Ansteuerung des Rücklaufventils zum Testen der Komponente 2
      OUT_V_Testen_K3 : Bool;   // Ansteuerung des Rücklaufventils zum Testen der Komponente 3
      OUT_V_Testen_K4 : Bool;   // Ansteuerung des Rücklaufventils zum Testen der Komponente 4
   END_VAR
   VAR_IN_OUT
      IO_Status : "UDT115_Test";   // Speichern der Testfunktions- Zustände für das Programm
   END_VAR
   VAR_TEMP
      Temp_IO_Status : "UDT115_Test";   // Temporärer Testfunktions- Status für die interne Bearbeitung des Bausteins
      ERROR_CODE : Int;   // Störungszustand der Systemfunktion "BLKMOV" Blockmove
      Anyzeiger : ANY;   // Zeiger zum Kopieren der Bereiche "IO_Status" und "Temp_IO_Status"
      Lampenansteuerung : Bool;   // Zwischenmerker für die Ansteuerung der Testanzeigen
   END_VAR
BEGIN

REGION Network 1: Gesicherte Daten einbinden
         LAR1;
         L;
         LAR2;
   //
         L     16#1002;  // Bytes
         T     W[AR1, P#0.0];
         L     2;  // Anzahl Bytes
         T     W[AR1, P#2.0];
         L     W[AR2, P#0.0];  // Baustein Nr.
         T     W[AR1, P#4.0];
         L     D[AR2, P#2.0];  // Datenanfang
         T     D[AR1, P#6.0];
   //
         CALL  BLKMOV
         ( SRCBLK  := #Anyzeiger,
           RET_VAL := #ERROR_CODE,
           DSTBLK  := #Temp_IO_Status
         );
   //
END_REGION

REGION Network 2
         ON    #IN_Betriebsart_Testen;
         O     #IN_Imp_Zyklus_Ende;
         ON    #IN_Stop_Testen;
         ON    #IN_Zyklus_Freigabe;
         JC    nTes;
   //
         O     #IN_Zyklus_Schuss_laeuft;
         O     #IN_Zyklus_KLZ2_u_ff;
         JC    Shot;
   //
         A     #IN_Start_Testen_K1;
         S     #Temp_IO_Status.Test_K1;
   //
         A     #IN_Start_Testen_K2;
         S     #Temp_IO_Status.Test_K2;
   //
         A     #IN_Start_Testen_K3;
         S     #Temp_IO_Status.Test_K3;
   //
         A     #IN_Start_Testen_K4;
         S     #Temp_IO_Status.Test_K4;
   //
         O     #Temp_IO_Status.Test_K1;
         O     #Temp_IO_Status.Test_K2;
         O     #Temp_IO_Status.Test_K3;
         O     #Temp_IO_Status.Test_K4;
         A     #IN_Zyklus_Freigabe;
         AN    #IN_Zyklus_laeuft;
         S     #Temp_IO_Status.Start_to_Cycle;
         S     #Temp_IO_Status.Test_runs;
   //
         A     #IN_Zyklus_laeuft;
         R     #Temp_IO_Status.Start_to_Cycle;
   //
   Shot: NOP   0;
   //
         A     #IN_Zyklus_Schuss_laeuft;
         A     #IN_Betriebsart_Betrieb;
         A     #Temp_IO_Status.Test_K1;
         =     #OUT_V_Testen_K1;
   //
         A     #IN_Zyklus_Schuss_laeuft;
         A     #IN_Betriebsart_Betrieb;
         A     #Temp_IO_Status.Test_K2;
         =     #OUT_V_Testen_K2;
   //
         A     #IN_Zyklus_Schuss_laeuft;
         A     #IN_Betriebsart_Betrieb;
         A     #Temp_IO_Status.Test_K3;
         =     #OUT_V_Testen_K3;
   //
         A     #IN_Zyklus_Schuss_laeuft;
         A     #IN_Betriebsart_Betrieb;
         A     #Temp_IO_Status.Test_K4;
         =     #OUT_V_Testen_K4;
   //
         ON    #Temp_IO_Status.Test_runs;
         O     #Temp_IO_Status.Start_to_Cycle;
         O     #IN_Zyklus_laeuft;
         AN    #IN_Stoerung_Gruppe_1;
         A     #IN_Stop_Testen;
         AN    #IN_Zyklus_KLZ2_u_ff;
         JC    Lamp;
   ///
   nTes: SET;
         A     #IN_Zyklus_laeuft;
         AN    #IN_Zyklus_KLZ2_u_ff;
         A     #Temp_IO_Status.Test_runs;
         =     #Temp_IO_Status.Stop_to_Cycle;
         SET;
         R     #Temp_IO_Status.Test_K1;
         R     #Temp_IO_Status.Test_K2;
         R     #Temp_IO_Status.Test_K3;
         R     #Temp_IO_Status.Test_K4;
         R     #Temp_IO_Status.Test_runs;
         R     #Temp_IO_Status.Start_to_Cycle;
         R     #OUT_V_Testen_K1;
         R     #OUT_V_Testen_K2;
         R     #OUT_V_Testen_K3;
         R     #OUT_V_Testen_K4;
END_REGION

REGION Network 3: Lampenansteuerung
   Lamp: A     #IN_Betriebsart_Testen;
         A     #IN_Zyklus_Freigabe;
         AN    #IN_Zyklus_laeuft;
         AN    #Temp_IO_Status.Test_runs;
         O;
         A     #IN_Betriebsart_Testen;
         A     #IN_Zyklus_laeuft;
         AN    #IN_Zyklus_Schuss_laeuft;
         A     #Temp_IO_Status.Test_runs;
         A     "Flag_01_000_Hertz";
         O;
         A     #IN_Betriebsart_Testen;
         A     #IN_Zyklus_laeuft;
         A     #IN_Zyklus_Schuss_laeuft;
         A     #Temp_IO_Status.Test_runs;
         A     "Flag_05_000_Hertz";
         O     #IN_Lampentest;
         =     #Lampenansteuerung;
   //
         ON    #Temp_IO_Status.Test_runs;
         O     #Temp_IO_Status.Test_K1;
         A     #Lampenansteuerung;
         =     #OUT_H_Testen_K1;
   //
         ON    #Temp_IO_Status.Test_runs;
         O     #Temp_IO_Status.Test_K2;
         A     #Lampenansteuerung;
         =     #OUT_H_Testen_K2;
   //
         ON    #Temp_IO_Status.Test_runs;
         O     #Temp_IO_Status.Test_K3;
         A     #Lampenansteuerung;
         =     #OUT_H_Testen_K3;
   //
         ON    #Temp_IO_Status.Test_runs;
         O     #Temp_IO_Status.Test_K4;
         A     #Lampenansteuerung;
         =     #OUT_H_Testen_K4;
END_REGION

REGION Network 4: Daten sichern
         CALL  BLKMOV
         ( SRCBLK  := #Temp_IO_Status,
           RET_VAL := #ERROR_CODE,
           DSTBLK  := #Anyzeiger
         );
   //
END_REGION
END_FUNCTION

